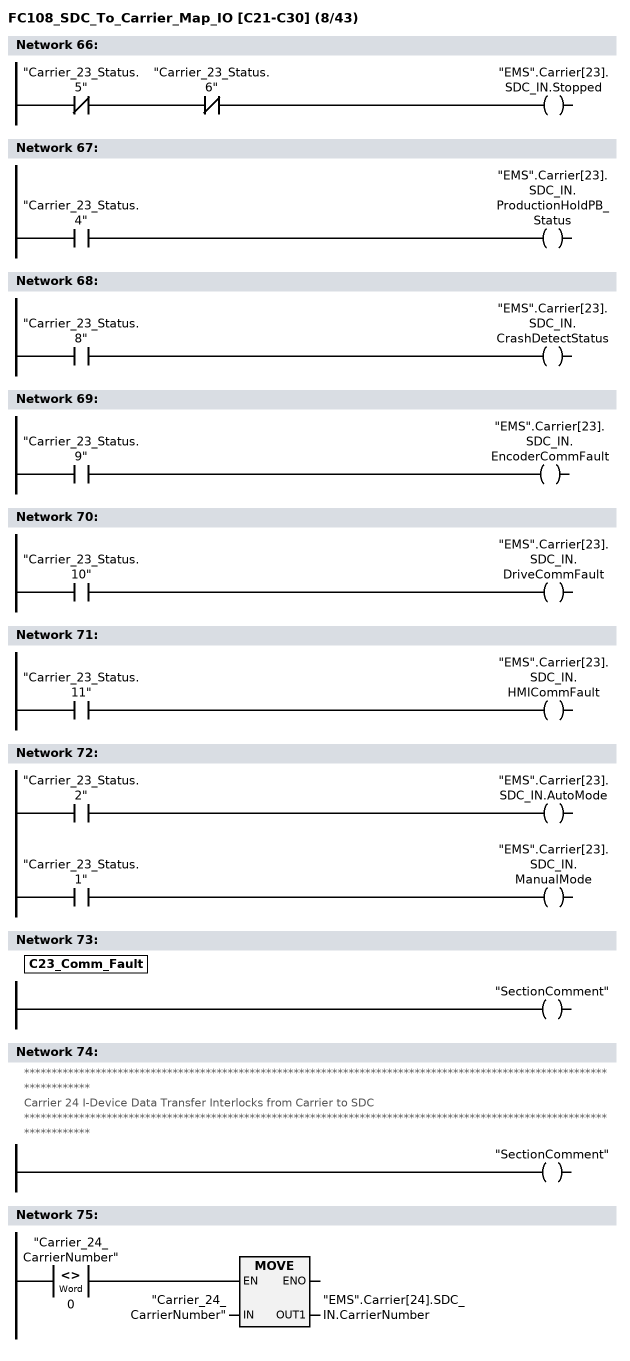
   RUNG wire#powerrail
      I_Contact( "Carrier_23_Status.5" )
      I_Contact( "Carrier_23_Status.6" )
      Coil( "EMS".Carrier[23].SDC_IN.Stopped )
   END_RUNG
   // the same network as SCL:
   "EMS".Carrier[23].SDC_IN.Stopped := NOT "Carrier_23_Status.5" AND NOT "Carrier_23_Status.6";
END_REGION

REGION Network 67
   RUNG wire#powerrail
      Contact( "Carrier_23_Status.4" )
      Coil( "EMS".Carrier[23].SDC_IN.ProductionHoldPB_Status )
   END_RUNG
   // the same network as SCL:
   "EMS".Carrier[23].SDC_IN.ProductionHoldPB_Status := "Carrier_23_Status.4";
END_REGION

REGION Network 68
   RUNG wire#powerrail
      Contact( "Carrier_23_Status.8" )
      Coil( "EMS".Carrier[23].SDC_IN.CrashDetectStatus )
   END_RUNG
   // the same network as SCL:
   "EMS".Carrier[23].SDC_IN.CrashDetectStatus := "Carrier_23_Status.8";
END_REGION

REGION Network 69
   RUNG wire#powerrail
      Contact( "Carrier_23_Status.9" )
      Coil( "EMS".Carrier[23].SDC_IN.EncoderCommFault )
   END_RUNG
   // the same network as SCL:
   "EMS".Carrier[23].SDC_IN.EncoderCommFault := "Carrier_23_Status.9";
END_REGION

REGION Network 70
   RUNG wire#powerrail
      Contact( "Carrier_23_Status.10" )
      Coil( "EMS".Carrier[23].SDC_IN.DriveCommFault )
   END_RUNG
   // the same network as SCL:
   "EMS".Carrier[23].SDC_IN.DriveCommFault := "Carrier_23_Status.10";
END_REGION

REGION Network 71
   RUNG wire#powerrail
      Contact( "Carrier_23_Status.11" )
      Coil( "EMS".Carrier[23].SDC_IN.HMICommFault )
   END_RUNG
   // the same network as SCL:
   "EMS".Carrier[23].SDC_IN.HMICommFault := "Carrier_23_Status.11";
END_REGION

REGION Network 72
   RUNG wire#powerrail
      Contact( "Carrier_23_Status.2" )
      Coil( "EMS".Carrier[23].SDC_IN.AutoMode )
   END_RUNG
   RUNG wire#powerrail
      Contact( "Carrier_23_Status.1" )
      Coil( "EMS".Carrier[23].SDC_IN.ManualMode )
   END_RUNG
   // the same network as SCL:
   "EMS".Carrier[23].SDC_IN.AutoMode := "Carrier_23_Status.2";
   "EMS".Carrier[23].SDC_IN.ManualMode := "Carrier_23_Status.1";
END_REGION

REGION Network 73
   Label( C23_Comm_Fault )
   RUNG wire#powerrail
      Coil( "SectionComment" )
   END_RUNG
   // the same network as SCL:
   C23_Comm_Fault:
   "SectionComment" := TRUE;
END_REGION

REGION Network 74
   // **********************************************************************************************************************
   // 
   // Carrier 24 I-Device Data Transfer Interlocks from Carrier to SDC
   // 
   // **********************************************************************************************************************
   RUNG wire#powerrail
      Coil( "SectionComment" )
   END_RUNG
   // the same network as SCL:
   "SectionComment" := TRUE;
END_REGION

REGION Network 75
   RUNG wire#powerrail
      { S7_Templates := "SrcType := Word" } NE_Contact(in1 := "Carrier_24_CarrierNumber", in2 := 0)
      Move(in := "Carrier_24_CarrierNumber", out1 => "EMS".Carrier[24].SDC_IN.CarrierNumber)
   END_RUNG
   // the same network as SCL:
   IF "Carrier_24_CarrierNumber" <> 0 THEN
       "EMS".Carrier[24].SDC_IN.CarrierNumber := "Carrier_24_CarrierNumber";
   END_IF;
END_REGION

REGION Network 76
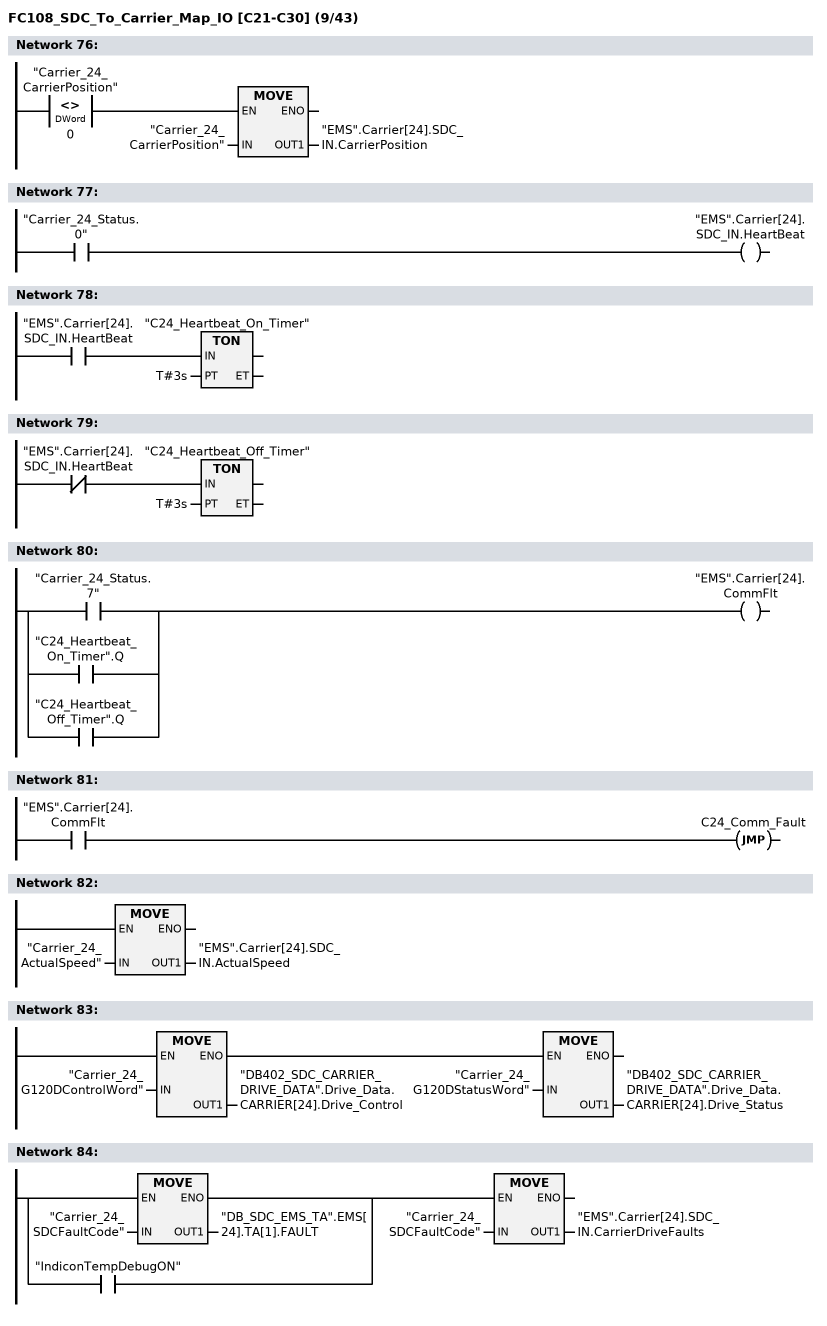
   RUNG wire#powerrail
      { S7_Templates := "SrcType := DWord" } NE_Contact(in1 := "Carrier_24_CarrierPosition", in2 := 0)
      Move(in := "Carrier_24_CarrierPosition", out1 => "EMS".Carrier[24].SDC_IN.CarrierPosition)
   END_RUNG
   // the same network as SCL:
   IF "Carrier_24_CarrierPosition" <> 0 THEN
       "EMS".Carrier[24].SDC_IN.CarrierPosition := "Carrier_24_CarrierPosition";
   END_IF;
END_REGION

REGION Network 77
   RUNG wire#powerrail
      Contact( "Carrier_24_Status.0" )
      Coil( "EMS".Carrier[24].SDC_IN.HeartBeat )
   END_RUNG
   // the same network as SCL:
   "EMS".Carrier[24].SDC_IN.HeartBeat := "Carrier_24_Status.0";
END_REGION

REGION Network 78
   "C24_Heartbeat_On_Timer".TON(IN := "EMS".Carrier[24].SDC_IN.HeartBeat, PT := T#3s);
END_REGION

REGION Network 79
   "C24_Heartbeat_Off_Timer".TON(IN := NOT "EMS".Carrier[24].SDC_IN.HeartBeat, PT := T#3s);
END_REGION

REGION Network 80
   RUNG wire#powerrail
      Contact( "Carrier_24_Status.7" )
      wire#w1
      Coil( "EMS".Carrier[24].CommFlt )
   END_RUNG
   RUNG wire#powerrail
      Contact( "C24_Heartbeat_On_Timer".Q )
   END_RUNG wire#w1
   RUNG wire#powerrail
      Contact( "C24_Heartbeat_Off_Timer".Q )
   END_RUNG wire#w1
   // the same network as SCL:
   "EMS".Carrier[24].CommFlt := "Carrier_24_Status.7" OR "C24_Heartbeat_On_Timer".Q OR "C24_Heartbeat_Off_Timer".Q;
END_REGION

REGION Network 81
   RUNG wire#powerrail
      Contact( "EMS".Carrier[24].CommFlt )
      JumpCoil( C24_Comm_Fault )
   END_RUNG
   // the same network as SCL:
   IF "EMS".Carrier[24].CommFlt THEN GOTO C24_Comm_Fault; END_IF;
END_REGION

REGION Network 82
   RUNG wire#powerrail
      Move(in := "Carrier_24_ActualSpeed", out1 => "EMS".Carrier[24].SDC_IN.ActualSpeed)
   END_RUNG
   // the same network as SCL:
   "EMS".Carrier[24].SDC_IN.ActualSpeed := "Carrier_24_ActualSpeed";
END_REGION

REGION Network 83
   RUNG wire#powerrail
      Move(in := "Carrier_24_G120DControlWord", out1 => "DB402_SDC_CARRIER_DRIVE_DATA".Drive_Data.CARRIER[24].Drive_Control)
      Move(in := "Carrier_24_G120DStatusWord", out1 => "DB402_SDC_CARRIER_DRIVE_DATA".Drive_Data.CARRIER[24].Drive_Status)
   END_RUNG
   // the same network as SCL:
   "DB402_SDC_CARRIER_DRIVE_DATA".Drive_Data.CARRIER[24].Drive_Control := "Carrier_24_G120DControlWord";
   "DB402_SDC_CARRIER_DRIVE_DATA".Drive_Data.CARRIER[24].Drive_Status := "Carrier_24_G120DStatusWord";
END_REGION

REGION Network 84
   RUNG wire#powerrail
      Move(in := "Carrier_24_SDCFaultCode", out1 => "DB_SDC_EMS_TA".EMS[24].TA[1].FAULT)
      wire#w1
      Move(in := "Carrier_24_SDCFaultCode", out1 => "EMS".Carrier[24].SDC_IN.CarrierDriveFaults)
   END_RUNG
   RUNG wire#powerrail
      Contact( "IndiconTempDebugON" )
   END_RUNG wire#w1
   // the same network as SCL:
   "DB_SDC_EMS_TA".EMS[24].TA[1].FAULT := "Carrier_24_SDCFaultCode";
   IF TRUE OR "IndiconTempDebugON" THEN
       "EMS".Carrier[24].SDC_IN.CarrierDriveFaults := "Carrier_24_SDCFaultCode";
   END_IF;
END_REGION

REGION Network 85
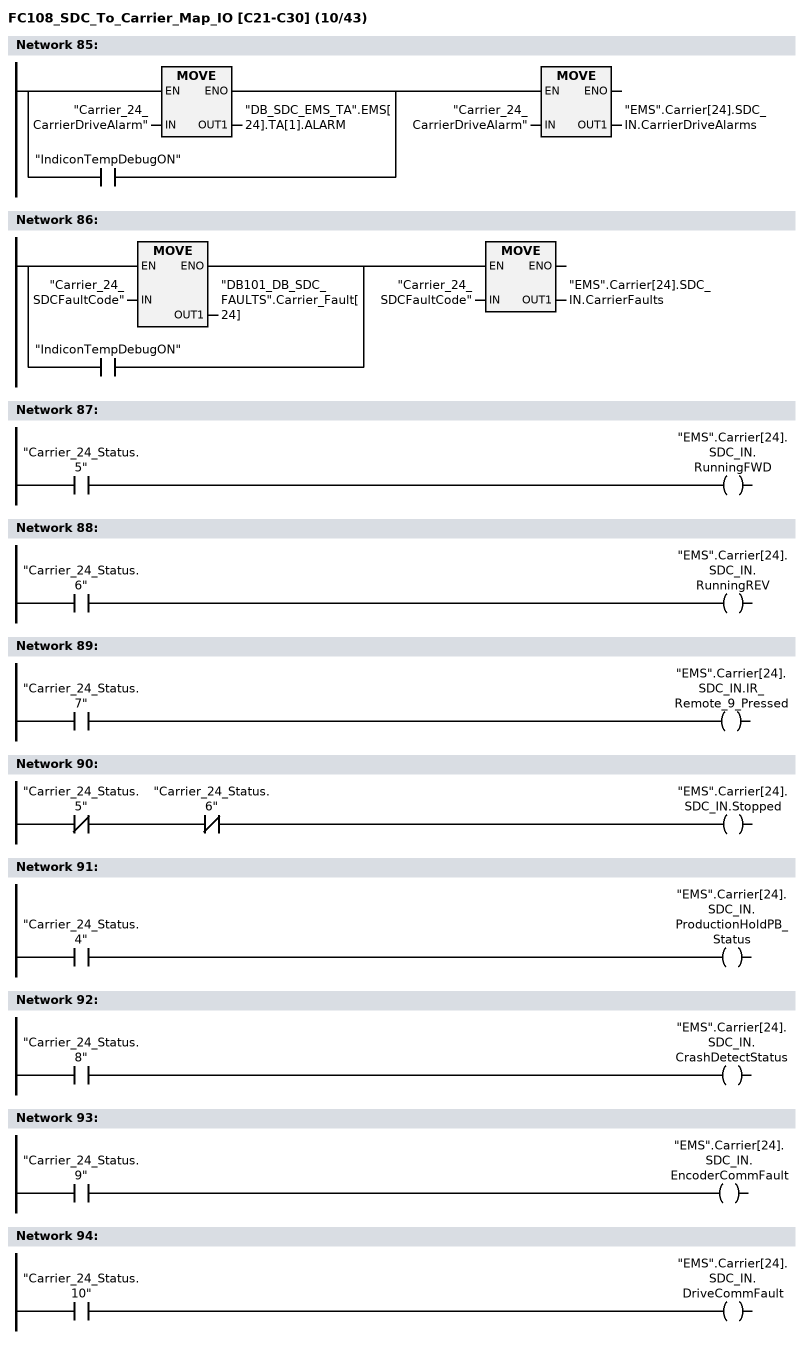
   RUNG wire#powerrail
      Move(in := "Carrier_24_CarrierDriveAlarm", out1 => "DB_SDC_EMS_TA".EMS[24].TA[1].ALARM)
      wire#w1
      Move(in := "Carrier_24_CarrierDriveAlarm", out1 => "EMS".Carrier[24].SDC_IN.CarrierDriveAlarms)
   END_RUNG
   RUNG wire#powerrail
      Contact( "IndiconTempDebugON" )
   END_RUNG wire#w1
   // the same network as SCL:
   "DB_SDC_EMS_TA".EMS[24].TA[1].ALARM := "Carrier_24_CarrierDriveAlarm";
   IF TRUE OR "IndiconTempDebugON" THEN
       "EMS".Carrier[24].SDC_IN.CarrierDriveAlarms := "Carrier_24_CarrierDriveAlarm";
   END_IF;
END_REGION

REGION Network 86
   RUNG wire#powerrail
      Move(in := "Carrier_24_SDCFaultCode", out1 => "DB101_DB_SDC_FAULTS".Carrier_Fault[24])
      wire#w1
      Move(in := "Carrier_24_SDCFaultCode", out1 => "EMS".Carrier[24].SDC_IN.CarrierFaults)
   END_RUNG
   RUNG wire#powerrail
      Contact( "IndiconTempDebugON" )
   END_RUNG wire#w1
   // the same network as SCL:
   "DB101_DB_SDC_FAULTS".Carrier_Fault[24] := "Carrier_24_SDCFaultCode";
   IF TRUE OR "IndiconTempDebugON" THEN
       "EMS".Carrier[24].SDC_IN.CarrierFaults := "Carrier_24_SDCFaultCode";
   END_IF;
END_REGION

REGION Network 87
   RUNG wire#powerrail
      Contact( "Carrier_24_Status.5" )
      Coil( "EMS".Carrier[24].SDC_IN.RunningFWD )
   END_RUNG
   // the same network as SCL:
   "EMS".Carrier[24].SDC_IN.RunningFWD := "Carrier_24_Status.5";
END_REGION

REGION Network 88
   RUNG wire#powerrail
      Contact( "Carrier_24_Status.6" )
      Coil( "EMS".Carrier[24].SDC_IN.RunningREV )
   END_RUNG
   // the same network as SCL:
   "EMS".Carrier[24].SDC_IN.RunningREV := "Carrier_24_Status.6";
END_REGION

REGION Network 89
   RUNG wire#powerrail
      Contact( "Carrier_24_Status.7" )
      Coil( "EMS".Carrier[24].SDC_IN.IR_Remote_9_Pressed )
   END_RUNG
   // the same network as SCL:
   "EMS".Carrier[24].SDC_IN.IR_Remote_9_Pressed := "Carrier_24_Status.7";
END_REGION

REGION Network 90
   RUNG wire#powerrail
      I_Contact( "Carrier_24_Status.5" )
      I_Contact( "Carrier_24_Status.6" )
      Coil( "EMS".Carrier[24].SDC_IN.Stopped )
   END_RUNG
   // the same network as SCL:
   "EMS".Carrier[24].SDC_IN.Stopped := NOT "Carrier_24_Status.5" AND NOT "Carrier_24_Status.6";
END_REGION

REGION Network 91
   RUNG wire#powerrail
      Contact( "Carrier_24_Status.4" )
      Coil( "EMS".Carrier[24].SDC_IN.ProductionHoldPB_Status )
   END_RUNG
   // the same network as SCL:
   "EMS".Carrier[24].SDC_IN.ProductionHoldPB_Status := "Carrier_24_Status.4";
END_REGION

REGION Network 92
   RUNG wire#powerrail
      Contact( "Carrier_24_Status.8" )
      Coil( "EMS".Carrier[24].SDC_IN.CrashDetectStatus )
   END_RUNG
   // the same network as SCL:
   "EMS".Carrier[24].SDC_IN.CrashDetectStatus := "Carrier_24_Status.8";
END_REGION

REGION Network 93
   RUNG wire#powerrail
      Contact( "Carrier_24_Status.9" )
      Coil( "EMS".Carrier[24].SDC_IN.EncoderCommFault )
   END_RUNG
   // the same network as SCL:
   "EMS".Carrier[24].SDC_IN.EncoderCommFault := "Carrier_24_Status.9";
END_REGION

REGION Network 94
   RUNG wire#powerrail
      Contact( "Carrier_24_Status.10" )
      Coil( "EMS".Carrier[24].SDC_IN.DriveCommFault )
   END_RUNG
   // the same network as SCL:
   "EMS".Carrier[24].SDC_IN.DriveCommFault := "Carrier_24_Status.10";
END_REGION

REGION Network 95
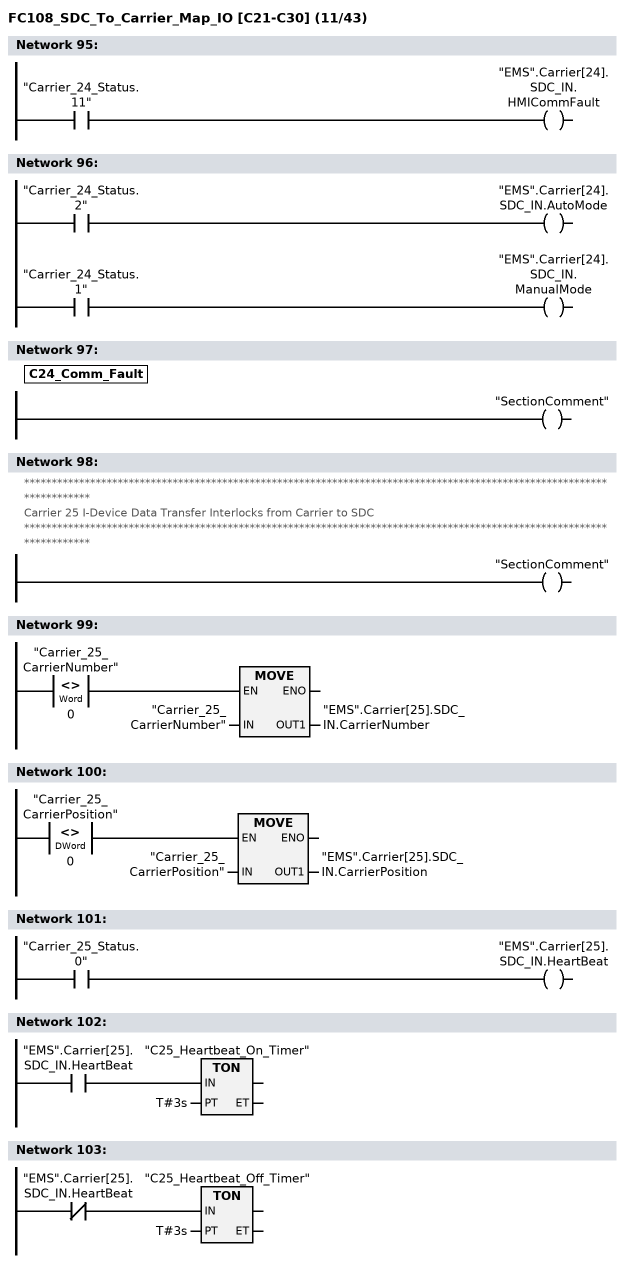
   RUNG wire#powerrail
      Contact( "Carrier_24_Status.11" )
      Coil( "EMS".Carrier[24].SDC_IN.HMICommFault )
   END_RUNG
   // the same network as SCL:
   "EMS".Carrier[24].SDC_IN.HMICommFault := "Carrier_24_Status.11";
END_REGION

REGION Network 96
   RUNG wire#powerrail
      Contact( "Carrier_24_Status.2" )
      Coil( "EMS".Carrier[24].SDC_IN.AutoMode )
   END_RUNG
   RUNG wire#powerrail
      Contact( "Carrier_24_Status.1" )
      Coil( "EMS".Carrier[24].SDC_IN.ManualMode )
   END_RUNG
   // the same network as SCL:
   "EMS".Carrier[24].SDC_IN.AutoMode := "Carrier_24_Status.2";
   "EMS".Carrier[24].SDC_IN.ManualMode := "Carrier_24_Status.1";
END_REGION

REGION Network 97
   Label( C24_Comm_Fault )
   RUNG wire#powerrail
      Coil( "SectionComment" )
   END_RUNG
   // the same network as SCL:
   C24_Comm_Fault:
   "SectionComment" := TRUE;
END_REGION

REGION Network 98
   // **********************************************************************************************************************
   // 
   // Carrier 25 I-Device Data Transfer Interlocks from Carrier to SDC
   // 
   // **********************************************************************************************************************
   RUNG wire#powerrail
      Coil( "SectionComment" )
   END_RUNG
   // the same network as SCL:
   "SectionComment" := TRUE;
END_REGION

REGION Network 99
   RUNG wire#powerrail
      { S7_Templates := "SrcType := Word" } NE_Contact(in1 := "Carrier_25_CarrierNumber", in2 := 0)
      Move(in := "Carrier_25_CarrierNumber", out1 => "EMS".Carrier[25].SDC_IN.CarrierNumber)
   END_RUNG
   // the same network as SCL:
   IF "Carrier_25_CarrierNumber" <> 0 THEN
       "EMS".Carrier[25].SDC_IN.CarrierNumber := "Carrier_25_CarrierNumber";
   END_IF;
END_REGION

REGION Network 100
   RUNG wire#powerrail
      { S7_Templates := "SrcType := DWord" } NE_Contact(in1 := "Carrier_25_CarrierPosition", in2 := 0)
      Move(in := "Carrier_25_CarrierPosition", out1 => "EMS".Carrier[25].SDC_IN.CarrierPosition)
   END_RUNG
   // the same network as SCL:
   IF "Carrier_25_CarrierPosition" <> 0 THEN
       "EMS".Carrier[25].SDC_IN.CarrierPosition := "Carrier_25_CarrierPosition";
   END_IF;
END_REGION

REGION Network 101
   RUNG wire#powerrail
      Contact( "Carrier_25_Status.0" )
      Coil( "EMS".Carrier[25].SDC_IN.HeartBeat )
   END_RUNG
   // the same network as SCL:
   "EMS".Carrier[25].SDC_IN.HeartBeat := "Carrier_25_Status.0";
END_REGION

REGION Network 102
   "C25_Heartbeat_On_Timer".TON(IN := "EMS".Carrier[25].SDC_IN.HeartBeat, PT := T#3s);
END_REGION

REGION Network 103
   "C25_Heartbeat_Off_Timer".TON(IN := NOT "EMS".Carrier[25].SDC_IN.HeartBeat, PT := T#3s);
END_REGION

REGION Network 104
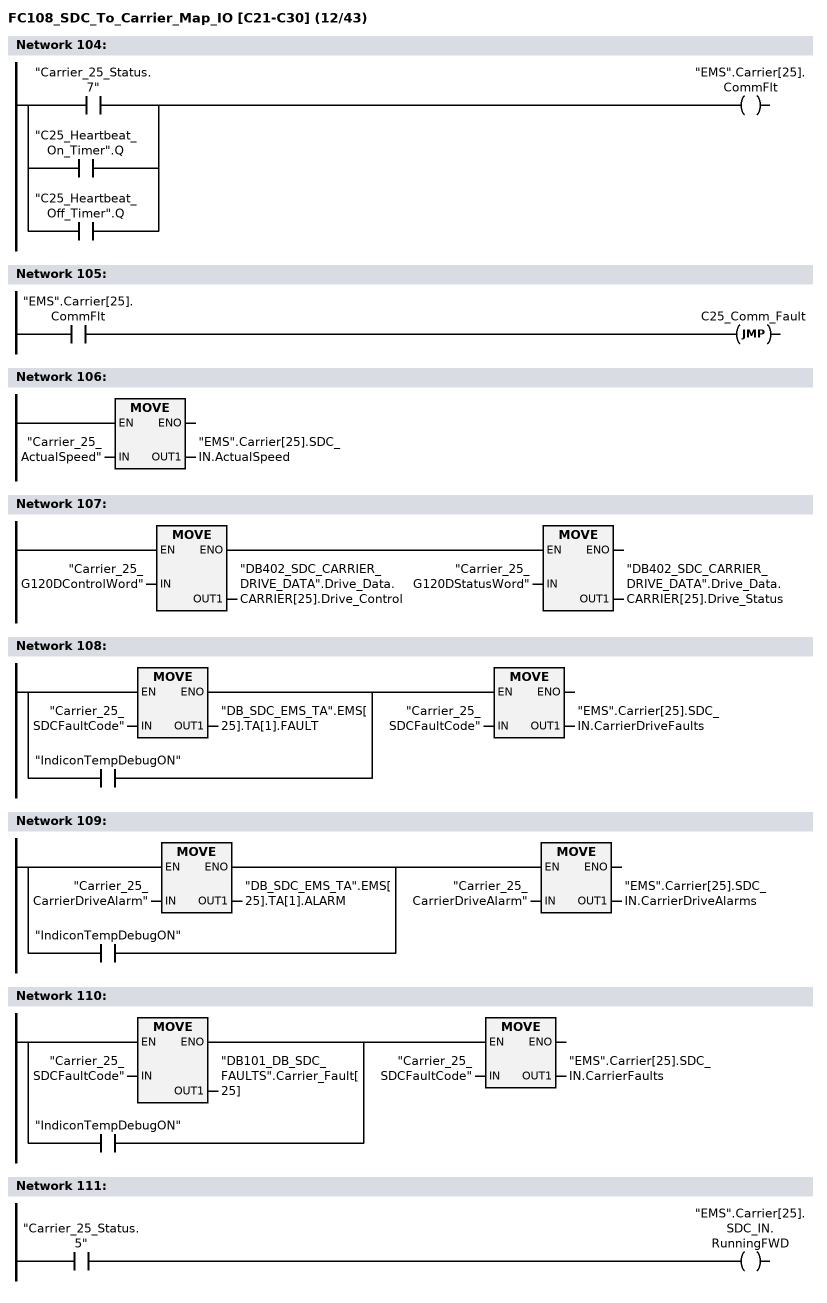
   RUNG wire#powerrail
      Contact( "Carrier_25_Status.7" )
      wire#w1
      Coil( "EMS".Carrier[25].CommFlt )
   END_RUNG
   RUNG wire#powerrail
      Contact( "C25_Heartbeat_On_Timer".Q )
   END_RUNG wire#w1
   RUNG wire#powerrail
      Contact( "C25_Heartbeat_Off_Timer".Q )
   END_RUNG wire#w1
   // the same network as SCL:
   "EMS".Carrier[25].CommFlt := "Carrier_25_Status.7" OR "C25_Heartbeat_On_Timer".Q OR "C25_Heartbeat_Off_Timer".Q;
END_REGION

REGION Network 105
   RUNG wire#powerrail
      Contact( "EMS".Carrier[25].CommFlt )
      JumpCoil( C25_Comm_Fault )
   END_RUNG
   // the same network as SCL:
   IF "EMS".Carrier[25].CommFlt THEN GOTO C25_Comm_Fault; END_IF;
END_REGION

REGION Network 106
   RUNG wire#powerrail
      Move(in := "Carrier_25_ActualSpeed", out1 => "EMS".Carrier[25].SDC_IN.ActualSpeed)
   END_RUNG
   // the same network as SCL:
   "EMS".Carrier[25].SDC_IN.ActualSpeed := "Carrier_25_ActualSpeed";
END_REGION

REGION Network 107
   RUNG wire#powerrail
      Move(in := "Carrier_25_G120DControlWord", out1 => "DB402_SDC_CARRIER_DRIVE_DATA".Drive_Data.CARRIER[25].Drive_Control)
      Move(in := "Carrier_25_G120DStatusWord", out1 => "DB402_SDC_CARRIER_DRIVE_DATA".Drive_Data.CARRIER[25].Drive_Status)
   END_RUNG
   // the same network as SCL:
   "DB402_SDC_CARRIER_DRIVE_DATA".Drive_Data.CARRIER[25].Drive_Control := "Carrier_25_G120DControlWord";
   "DB402_SDC_CARRIER_DRIVE_DATA".Drive_Data.CARRIER[25].Drive_Status := "Carrier_25_G120DStatusWord";
END_REGION

REGION Network 108
   RUNG wire#powerrail
      Move(in := "Carrier_25_SDCFaultCode", out1 => "DB_SDC_EMS_TA".EMS[25].TA[1].FAULT)
      wire#w1
      Move(in := "Carrier_25_SDCFaultCode", out1 => "EMS".Carrier[25].SDC_IN.CarrierDriveFaults)
   END_RUNG
   RUNG wire#powerrail
      Contact( "IndiconTempDebugON" )
   END_RUNG wire#w1
   // the same network as SCL:
   "DB_SDC_EMS_TA".EMS[25].TA[1].FAULT := "Carrier_25_SDCFaultCode";
   IF TRUE OR "IndiconTempDebugON" THEN
       "EMS".Carrier[25].SDC_IN.CarrierDriveFaults := "Carrier_25_SDCFaultCode";
   END_IF;
END_REGION

REGION Network 109
   RUNG wire#powerrail
      Move(in := "Carrier_25_CarrierDriveAlarm", out1 => "DB_SDC_EMS_TA".EMS[25].TA[1].ALARM)
      wire#w1
      Move(in := "Carrier_25_CarrierDriveAlarm", out1 => "EMS".Carrier[25].SDC_IN.CarrierDriveAlarms)
   END_RUNG
   RUNG wire#powerrail
      Contact( "IndiconTempDebugON" )
   END_RUNG wire#w1
   // the same network as SCL:
   "DB_SDC_EMS_TA".EMS[25].TA[1].ALARM := "Carrier_25_CarrierDriveAlarm";
   IF TRUE OR "IndiconTempDebugON" THEN
       "EMS".Carrier[25].SDC_IN.CarrierDriveAlarms := "Carrier_25_CarrierDriveAlarm";
   END_IF;
END_REGION

REGION Network 110
   RUNG wire#powerrail
      Move(in := "Carrier_25_SDCFaultCode", out1 => "DB101_DB_SDC_FAULTS".Carrier_Fault[25])
      wire#w1
      Move(in := "Carrier_25_SDCFaultCode", out1 => "EMS".Carrier[25].SDC_IN.CarrierFaults)
   END_RUNG
   RUNG wire#powerrail
      Contact( "IndiconTempDebugON" )
   END_RUNG wire#w1
   // the same network as SCL:
   "DB101_DB_SDC_FAULTS".Carrier_Fault[25] := "Carrier_25_SDCFaultCode";
   IF TRUE OR "IndiconTempDebugON" THEN
       "EMS".Carrier[25].SDC_IN.CarrierFaults := "Carrier_25_SDCFaultCode";
   END_IF;
END_REGION

REGION Network 111
   RUNG wire#powerrail
      Contact( "Carrier_25_Status.5" )
      Coil( "EMS".Carrier[25].SDC_IN.RunningFWD )
   END_RUNG
   // the same network as SCL:
   "EMS".Carrier[25].SDC_IN.RunningFWD := "Carrier_25_Status.5";
END_REGION

REGION Network 112
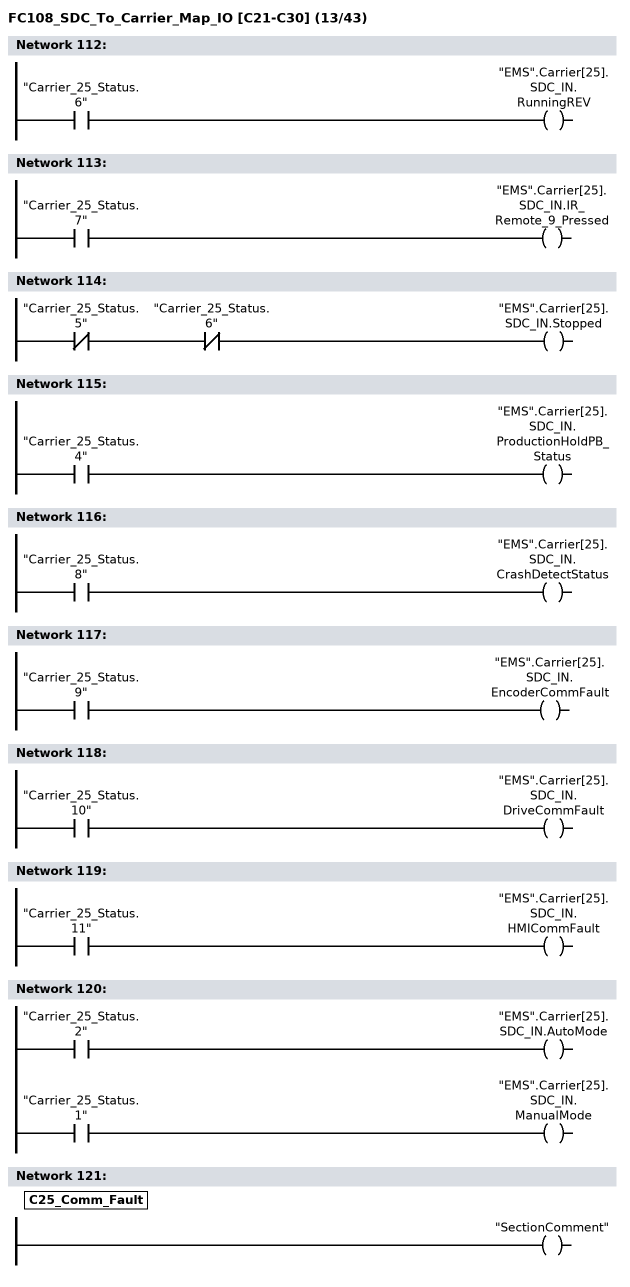
   RUNG wire#powerrail
      Contact( "Carrier_25_Status.6" )
      Coil( "EMS".Carrier[25].SDC_IN.RunningREV )
   END_RUNG
   // the same network as SCL:
   "EMS".Carrier[25].SDC_IN.RunningREV := "Carrier_25_Status.6";
END_REGION

REGION Network 113
   RUNG wire#powerrail
      Contact( "Carrier_25_Status.7" )
      Coil( "EMS".Carrier[25].SDC_IN.IR_Remote_9_Pressed )
   END_RUNG
   // the same network as SCL:
   "EMS".Carrier[25].SDC_IN.IR_Remote_9_Pressed := "Carrier_25_Status.7";
END_REGION

REGION Network 114
   RUNG wire#powerrail
      I_Contact( "Carrier_25_Status.5" )
      I_Contact( "Carrier_25_Status.6" )
      Coil( "EMS".Carrier[25].SDC_IN.Stopped )
   END_RUNG
   // the same network as SCL:
   "EMS".Carrier[25].SDC_IN.Stopped := NOT "Carrier_25_Status.5" AND NOT "Carrier_25_Status.6";
END_REGION

REGION Network 115
   RUNG wire#powerrail
      Contact( "Carrier_25_Status.4" )
      Coil( "EMS".Carrier[25].SDC_IN.ProductionHoldPB_Status )
   END_RUNG
   // the same network as SCL:
   "EMS".Carrier[25].SDC_IN.ProductionHoldPB_Status := "Carrier_25_Status.4";
END_REGION

REGION Network 116
   RUNG wire#powerrail
      Contact( "Carrier_25_Status.8" )
      Coil( "EMS".Carrier[25].SDC_IN.CrashDetectStatus )
   END_RUNG
   // the same network as SCL:
   "EMS".Carrier[25].SDC_IN.CrashDetectStatus := "Carrier_25_Status.8";
END_REGION

REGION Network 117
   RUNG wire#powerrail
      Contact( "Carrier_25_Status.9" )
      Coil( "EMS".Carrier[25].SDC_IN.EncoderCommFault )
   END_RUNG
   // the same network as SCL:
   "EMS".Carrier[25].SDC_IN.EncoderCommFault := "Carrier_25_Status.9";
END_REGION

REGION Network 118
   RUNG wire#powerrail
      Contact( "Carrier_25_Status.10" )
      Coil( "EMS".Carrier[25].SDC_IN.DriveCommFault )
   END_RUNG
   // the same network as SCL:
   "EMS".Carrier[25].SDC_IN.DriveCommFault := "Carrier_25_Status.10";
END_REGION

REGION Network 119
   RUNG wire#powerrail
      Contact( "Carrier_25_Status.11" )
      Coil( "EMS".Carrier[25].SDC_IN.HMICommFault )
   END_RUNG
   // the same network as SCL:
   "EMS".Carrier[25].SDC_IN.HMICommFault := "Carrier_25_Status.11";
END_REGION

REGION Network 120
   RUNG wire#powerrail
      Contact( "Carrier_25_Status.2" )
      Coil( "EMS".Carrier[25].SDC_IN.AutoMode )
   END_RUNG
   RUNG wire#powerrail
      Contact( "Carrier_25_Status.1" )
      Coil( "EMS".Carrier[25].SDC_IN.ManualMode )
   END_RUNG
   // the same network as SCL:
   "EMS".Carrier[25].SDC_IN.AutoMode := "Carrier_25_Status.2";
   "EMS".Carrier[25].SDC_IN.ManualMode := "Carrier_25_Status.1";
END_REGION

REGION Network 121
   Label( C25_Comm_Fault )
   RUNG wire#powerrail
      Coil( "SectionComment" )
   END_RUNG
   // the same network as SCL:
   C25_Comm_Fault:
   "SectionComment" := TRUE;
END_REGION

REGION Network 122
   // **********************************************************************************************************************
   // 
   // Carrier 26 I-Device Data Transfer Interlocks from Carrier to SDC
   // 
   // **********************************************************************************************************************
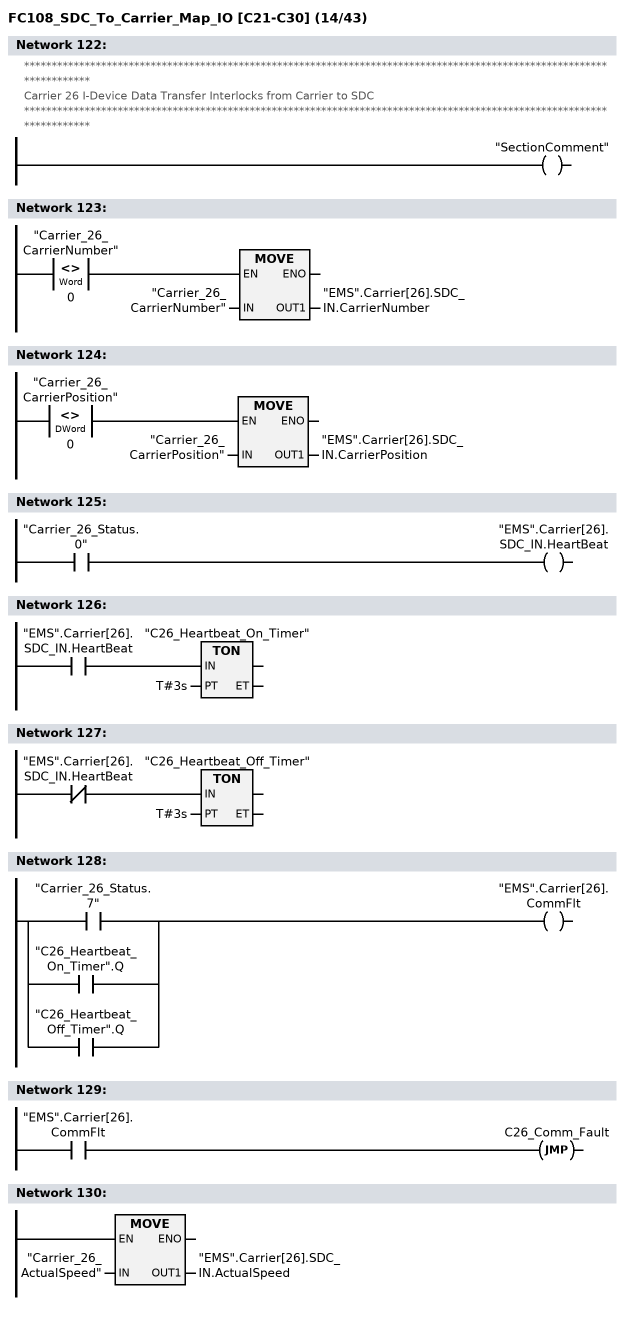
   RUNG wire#powerrail
      Coil( "SectionComment" )
   END_RUNG
   // the same network as SCL:
   "SectionComment" := TRUE;
END_REGION

REGION Network 123
   RUNG wire#powerrail
      { S7_Templates := "SrcType := Word" } NE_Contact(in1 := "Carrier_26_CarrierNumber", in2 := 0)
      Move(in := "Carrier_26_CarrierNumber", out1 => "EMS".Carrier[26].SDC_IN.CarrierNumber)
   END_RUNG
   // the same network as SCL:
   IF "Carrier_26_CarrierNumber" <> 0 THEN
       "EMS".Carrier[26].SDC_IN.CarrierNumber := "Carrier_26_CarrierNumber";
   END_IF;
END_REGION

REGION Network 124
   RUNG wire#powerrail
      { S7_Templates := "SrcType := DWord" } NE_Contact(in1 := "Carrier_26_CarrierPosition", in2 := 0)
      Move(in := "Carrier_26_CarrierPosition", out1 => "EMS".Carrier[26].SDC_IN.CarrierPosition)
   END_RUNG
   // the same network as SCL:
   IF "Carrier_26_CarrierPosition" <> 0 THEN
       "EMS".Carrier[26].SDC_IN.CarrierPosition := "Carrier_26_CarrierPosition";
   END_IF;
END_REGION

REGION Network 125
   RUNG wire#powerrail
      Contact( "Carrier_26_Status.0" )
      Coil( "EMS".Carrier[26].SDC_IN.HeartBeat )
   END_RUNG
   // the same network as SCL:
   "EMS".Carrier[26].SDC_IN.HeartBeat := "Carrier_26_Status.0";
END_REGION

REGION Network 126
   "C26_Heartbeat_On_Timer".TON(IN := "EMS".Carrier[26].SDC_IN.HeartBeat, PT := T#3s);
END_REGION

REGION Network 127
   "C26_Heartbeat_Off_Timer".TON(IN := NOT "EMS".Carrier[26].SDC_IN.HeartBeat, PT := T#3s);
END_REGION

REGION Network 128
   RUNG wire#powerrail
      Contact( "Carrier_26_Status.7" )
      wire#w1
      Coil( "EMS".Carrier[26].CommFlt )
   END_RUNG
   RUNG wire#powerrail
      Contact( "C26_Heartbeat_On_Timer".Q )
   END_RUNG wire#w1
   RUNG wire#powerrail
      Contact( "C26_Heartbeat_Off_Timer".Q )
   END_RUNG wire#w1
   // the same network as SCL:
   "EMS".Carrier[26].CommFlt := "Carrier_26_Status.7" OR "C26_Heartbeat_On_Timer".Q OR "C26_Heartbeat_Off_Timer".Q;
END_REGION

REGION Network 129
   RUNG wire#powerrail
      Contact( "EMS".Carrier[26].CommFlt )
      JumpCoil( C26_Comm_Fault )
   END_RUNG
   // the same network as SCL:
   IF "EMS".Carrier[26].CommFlt THEN GOTO C26_Comm_Fault; END_IF;
END_REGION

REGION Network 130
   RUNG wire#powerrail
      Move(in := "Carrier_26_ActualSpeed", out1 => "EMS".Carrier[26].SDC_IN.ActualSpeed)
   END_RUNG
   // the same network as SCL:
   "EMS".Carrier[26].SDC_IN.ActualSpeed := "Carrier_26_ActualSpeed";
END_REGION

REGION Network 131
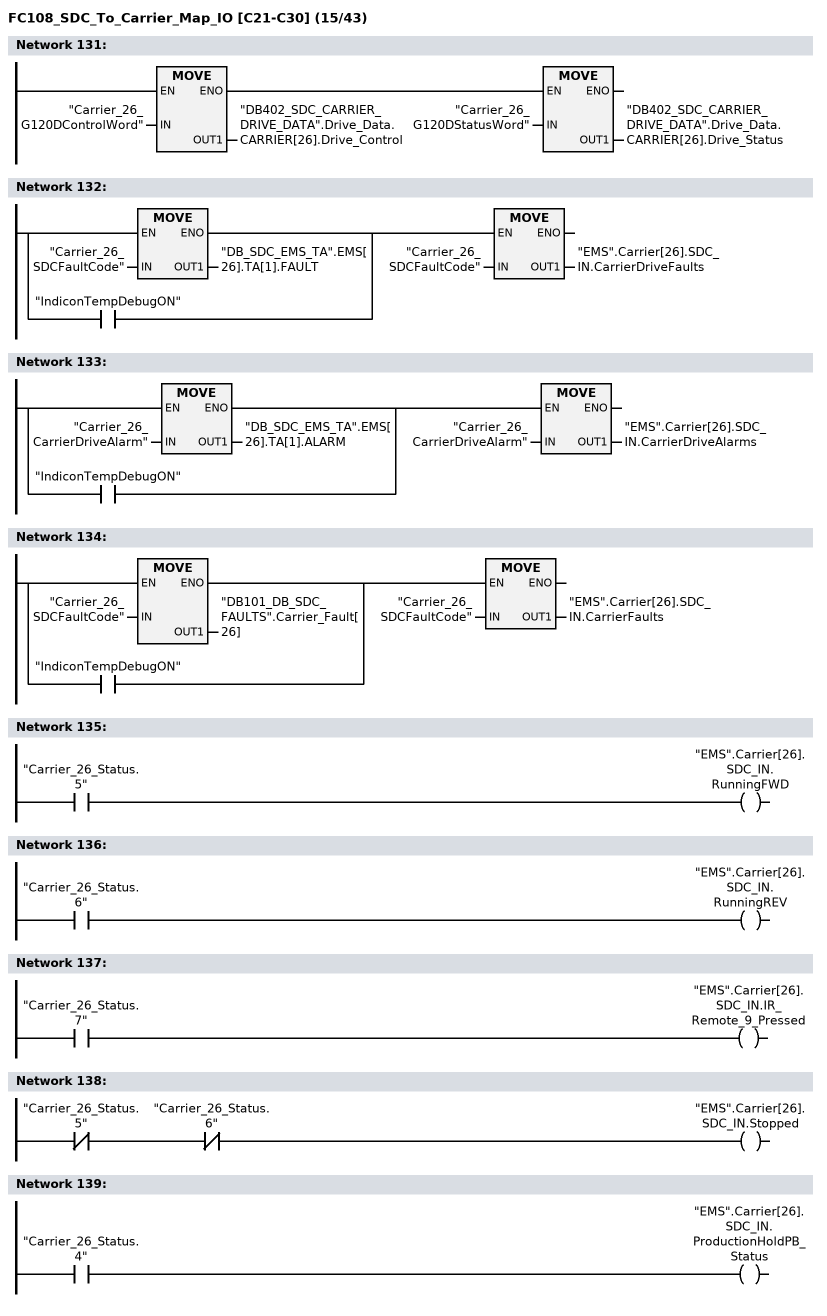
   RUNG wire#powerrail
      Move(in := "Carrier_26_G120DControlWord", out1 => "DB402_SDC_CARRIER_DRIVE_DATA".Drive_Data.CARRIER[26].Drive_Control)
      Move(in := "Carrier_26_G120DStatusWord", out1 => "DB402_SDC_CARRIER_DRIVE_DATA".Drive_Data.CARRIER[26].Drive_Status)
   END_RUNG
   // the same network as SCL:
   "DB402_SDC_CARRIER_DRIVE_DATA".Drive_Data.CARRIER[26].Drive_Control := "Carrier_26_G120DControlWord";
   "DB402_SDC_CARRIER_DRIVE_DATA".Drive_Data.CARRIER[26].Drive_Status := "Carrier_26_G120DStatusWord";
END_REGION

REGION Network 132
   RUNG wire#powerrail
      Move(in := "Carrier_26_SDCFaultCode", out1 => "DB_SDC_EMS_TA".EMS[26].TA[1].FAULT)
      wire#w1
      Move(in := "Carrier_26_SDCFaultCode", out1 => "EMS".Carrier[26].SDC_IN.CarrierDriveFaults)
   END_RUNG
   RUNG wire#powerrail
      Contact( "IndiconTempDebugON" )
   END_RUNG wire#w1
   // the same network as SCL:
   "DB_SDC_EMS_TA".EMS[26].TA[1].FAULT := "Carrier_26_SDCFaultCode";
   IF TRUE OR "IndiconTempDebugON" THEN
       "EMS".Carrier[26].SDC_IN.CarrierDriveFaults := "Carrier_26_SDCFaultCode";
   END_IF;
END_REGION

REGION Network 133
   RUNG wire#powerrail
      Move(in := "Carrier_26_CarrierDriveAlarm", out1 => "DB_SDC_EMS_TA".EMS[26].TA[1].ALARM)
      wire#w1
      Move(in := "Carrier_26_CarrierDriveAlarm", out1 => "EMS".Carrier[26].SDC_IN.CarrierDriveAlarms)
   END_RUNG
   RUNG wire#powerrail
      Contact( "IndiconTempDebugON" )
   END_RUNG wire#w1
   // the same network as SCL:
   "DB_SDC_EMS_TA".EMS[26].TA[1].ALARM := "Carrier_26_CarrierDriveAlarm";
   IF TRUE OR "IndiconTempDebugON" THEN
       "EMS".Carrier[26].SDC_IN.CarrierDriveAlarms := "Carrier_26_CarrierDriveAlarm";
   END_IF;
END_REGION

REGION Network 134
   RUNG wire#powerrail
      Move(in := "Carrier_26_SDCFaultCode", out1 => "DB101_DB_SDC_FAULTS".Carrier_Fault[26])
      wire#w1
      Move(in := "Carrier_26_SDCFaultCode", out1 => "EMS".Carrier[26].SDC_IN.CarrierFaults)
   END_RUNG
   RUNG wire#powerrail
      Contact( "IndiconTempDebugON" )
   END_RUNG wire#w1
   // the same network as SCL:
   "DB101_DB_SDC_FAULTS".Carrier_Fault[26] := "Carrier_26_SDCFaultCode";
   IF TRUE OR "IndiconTempDebugON" THEN
       "EMS".Carrier[26].SDC_IN.CarrierFaults := "Carrier_26_SDCFaultCode";
   END_IF;
END_REGION

REGION Network 135
   RUNG wire#powerrail
      Contact( "Carrier_26_Status.5" )
      Coil( "EMS".Carrier[26].SDC_IN.RunningFWD )
   END_RUNG
   // the same network as SCL:
   "EMS".Carrier[26].SDC_IN.RunningFWD := "Carrier_26_Status.5";
END_REGION

REGION Network 136
   RUNG wire#powerrail
      Contact( "Carrier_26_Status.6" )
      Coil( "EMS".Carrier[26].SDC_IN.RunningREV )
   END_RUNG
   // the same network as SCL:
   "EMS".Carrier[26].SDC_IN.RunningREV := "Carrier_26_Status.6";
END_REGION
